               IF NOT #statIsArrayFieldClosed THEN
                 //field wasn't close as no deeper hierarchy exist, therfore the normal close opeartion is invalid
                 //close now here
                 #statInfoToWrite := CONCAT(IN1 := CHAR_TO_STRING(#BRACES_CLOSE), IN2 := CHAR_TO_STRING(#COMMA));
                 #statStackIndex -= #DECREMENT_BY_ONE;
               ELSE //reset flag
                 #statIsArrayFieldClosed := FALSE;
               END_IF;
               //open object
               #statInfoToWrite := CONCAT(IN1 := #statInfoToWrite, IN2 := CHAR_TO_STRING(#BRACES_OPEN), IN3 := CHAR_TO_STRING(#WHITE_SPACE));
               //increase stack index and push closing elements on to it
               #statStackIndex += #INCREMENT_BY_ONE;
               #statStackIndexOpenElement[#statStackIndex] := #BRACES_CLOSE;
             END_IF;

             IF NOT (#statIsArrayOpen AND #statArrayName = #tree[#statIndexTreeArray].key)  THEN
               //write key not in case array is open and key is the same array name
               //this indicates simple array structure e.g "ArrayName":["ArrayValue1","ArrayValue2"]
               //write key -> "key":
               #statInfoToWrite := CONCAT(IN1 := #statInfoToWrite, IN2 := CHAR_TO_STRING(#QUTATIONMARK),
                                          IN3 := #tree[#statIndexTreeArray].key, IN4 := CHAR_TO_STRING(#QUTATIONMARK),
                                          IN5 := CHAR_TO_STRING(#COLON), IN6 := CHAR_TO_STRING(#WHITE_SPACE));

             END_IF;

             //Move to state Write
             #statFbState := #FB_STATE_WRITE_TO_JSON;
             //Set state, that should be executed after writing
             //move on to next state
             #statFbNextState := #FB_STATE_VALUE_TYPE;

           END_REGION NEXT_ELEMENT 

         #FB_STATE_VALUE_TYPE: // Depending on value type, write value
           REGION VALUE DEPENDECY OF TYPE
             CASE #tree[#statIndexTreeArray].type OF

               #OBJECT:
                 REGION OBJECT
                   //nothing to do when type is object just add line feed, { openning will occur with next depth
                   #statInfoToWrite := CONCAT(IN1 := #statInfoToWrite, IN2 := CHAR_TO_STRING(#BRACES_OPEN));
                   //increase stack index and push closing elements on to it
                   #statStackIndex += #INCREMENT_BY_ONE;
                   #statStackIndexOpenElement[#statStackIndex] := #BRACES_CLOSE;
                 END_REGION OBJECT

               #ARRAY:
                 REGION ARRAY

                   IF (NOT #statIsArrayOpen) THEN
                     #statIsFirstElement := TRUE;
                     #statIsArrayOpen := TRUE;
                     //set Name of Array
                     #statArrayName := #tree[#statIndexTreeArray].key;

                     #statInfoToWrite := CONCAT(IN1 := CHAR_TO_STRING(#BRACKETS_OPEN), IN2 := CHAR_TO_STRING(#WHITE_SPACE));
                     //increase stack index and push closing elements on to it
                     #statStackIndex += #INCREMENT_BY_ONE;
                     #statStackIndexOpenElement[#statStackIndex] := #BRACKETS_CLOSE;

                     //case for underlaying object structure in array, prevent depth of simple array to have leading {
                     //simple array always has arrayname as key
                     IF #tree[#statIndexTreeArray].depth < #tree[#statIndexTreeArray + #NEXT_INDEX].depth
                       AND #tree[#statIndexTreeArray+ #NEXT_INDEX].key <> #statArrayName THEN
                       //open object
                       #statInfoToWrite := CONCAT(IN1 := #statInfoToWrite, IN2 := CHAR_TO_STRING(#BRACES_OPEN));
                       //increase stack index and push closing elements on to it
                       #statStackIndex += #INCREMENT_BY_ONE;
                       #statStackIndexOpenElement[#statStackIndex] := #BRACES_CLOSE;
                     END_IF;

                   END_IF;

                   // //null indicating that it is array definition, array information is written sepe
                   // //otherwise write value as string - value enclosed with quotation mark 
                   // IF(#tree[#statIndexTreeArray].value <> #NULL) THEN
                   //   #statInfoToWrite := CONCAT(IN1 := #statInfoToWrite, IN2 := CHAR_TO_STRING(#QUTATIONMARK),
                   //                              IN3 := #tree[#statIndexTreeArray].value, IN4 := CHAR_TO_STRING(#QUTATIONMARK));
                   // END_IF;
                 END_REGION ARRAY 

               #STRING:
                 REGION STRING

                   //wirte value as string - value enclosed with quotation mark 
                   IF (#tree[#statIndexTreeArray].value <> #NULL) THEN
                     #statInfoToWrite := CONCAT(IN1 := #statInfoToWrite, IN2 := CHAR_TO_STRING(#QUTATIONMARK),
                                                IN3 := #tree[#statIndexTreeArray].value, IN4 := CHAR_TO_STRING(#QUTATIONMARK));

                   ELSE // empty value still needs "" otherwise syntax error
                     #statInfoToWrite := CONCAT(IN1 := #statInfoToWrite, IN2 := CHAR_TO_STRING(#QUTATIONMARK),
                                                IN3 := CHAR_TO_STRING(#QUTATIONMARK));
                   END_IF;
                 END_REGION STRING

               #NUMBER, #BOOLEAN:
                 REGION NUMBER_BOOLEAN
                   //wirte value as number or boolean - value enclosed without quotation mark 
                   IF (#tree[#statIndexTreeArray].value <> #NULL) THEN
                     #statInfoToWrite := CONCAT(IN1 := #statInfoToWrite,
                                                IN2 := #tree[#statIndexTreeArray].value);
                   END_IF;
                 END_REGION NUMBER_BOOLEAN

               ELSE // Undefined state in state machine reached
                 REGION UNDEFINED STATE
                   #statStatus := #ERR_UNDEFINED_STATE;
                 END_REGION UNDEFINED STATE          

             END_CASE;

             //Move to state Write
             #statFbState := #FB_STATE_WRITE_TO_JSON;

             //Set state, that should be executed after writing
             //move on to next state
             #statFbNextState := #FB_STATE_NEXT_ELEMENT;

             IF #statIsLastElement OR #tree[#statIndexTreeArray].depth > #tree[#statIndexTreeArray + #NEXT_INDEX].depth THEN
               //Next Element has lower depth, therefore Elements have to be closed
               #statFbNextState := #FB_STATE_CLOSE_STACK_ELEMENT;
             ELSIF #statIsLastElement OR #tree[#statIndexTreeArray].depth = #tree[#statIndexTreeArray + #NEXT_INDEX].depth AND  NOT #statIsFirstElement THEN
                #statInfoToWrite := CONCAT(IN1 := #statInfoToWrite,
                                           IN2 := CHAR_TO_STRING(#COMMA));
             END_IF;
             //#statInfoToWrite := CONCAT(IN1 := #statInfoToWrite, IN2 := CHAR_TO_STRING(#LINE_FEED));



             //increase tree index to access next element 
             #statIndexTreeArray += #INCREMENT_BY_ONE;

           END_REGION VALUE DEPENDECY OF TYPE

         #FB_STATE_WRITE_TO_JSON: // Write to Byte Array
           REGION WRITE TO JSON                
             //add information to json byte array
             IF ((INT_TO_UINT(LEN(#statInfoToWrite)) + #statIndexJsonByteArray) < #statJsonByteLen) THEN
               Strg_TO_Chars(Strg := #statInfoToWrite,
                             pChars := #statIndexJsonByteArray,
                             Cnt => #tempCntCharsAdded,
                             Chars := #jsonByteArray);


               #statInfoToWrite := #EMPTY;
               //move index of byte array 
               #statIndexJsonByteArray += #tempCntCharsAdded;
               //move to next state previously allocated
               #statFbState := #statFbNextState;
             ELSE // Error: Index out of bounds
               #statStatus := #ERR_JSON_OUT_OF_BOUNDS;
             END_IF;

             IF #statLastElementIsClosed THEN
               //writer has written last information and execution is done
               #statStatus := #STATUS_EXECUTION_FINISHED;
               //current index equals count/size of json byte array
               #statCount := #statIndexJsonByteArray;
             END_IF;
           END_REGION WRITE TO JSON

         #FB_STATE_CLOSE_STACK_ELEMENT: //Close Open Stack Elements
           REGION CLOSE ELEMENT FROM STACK
             //close element with syntax </key>

             IF #statStackIndex >= 0 THEN //more open elements available, not all elements are closed

               //statInfoToWrite --> } or ]
               #statInfoToWrite := CHAR_TO_STRING(#statStackIndexOpenElement[#statStackIndex]);

               IF #statInfoToWrite = #BRACKETS_CLOSE THEN
                 //reset flag
                 #statIsArrayOpen := FALSE;

                 //first array key is used to recognize,
                 //beginning of new array field reset here, so it can be check for emptiness
                 #statFirstArrayKey := '';
               END_IF;

               //pop element from stack 
               #statStackIndex -= SINT_TO_INT(#DECREMENT_BY_ONE);

               IF #statStackIndex >= 0 THEN //more open elements available, not all elements are closed
                 //look at current stack item depth, if next tree element has 
                 IF NOT #statIsLastElement AND #statStackIndex = #tree[#statIndexTreeArray].depth THEN
                   //move to next element
                   //write comma as JSON dictates same depth a divided by comma,
                   //here we move on to the next elment with the same depth
                   #statInfoToWrite := CONCAT(IN1:=  #statInfoToWrite, IN2:= CHAR_TO_STRING(#COMMA));

                   // //if Array is still open and the same lenght is reached,
                   // //new element in array, distinguish new entry with BRACES
                   IF #statIsArrayOpen THEN
                     #statInfoToWrite := CONCAT(IN1 := #statInfoToWrite, IN2 := CHAR_TO_STRING(#BRACES_CLOSE), IN3 := CHAR_TO_STRING(#COMMA));
                     //pop element from stack 
                     #statStackIndex -= SINT_TO_INT(#DECREMENT_BY_ONE);
                     #statIsArrayFieldClosed := TRUE;
                   //   #statInfoToWrite := CONCAT(IN1 := #statInfoToWrite, IN2 := CHAR_TO_STRING(#BRACES_OPEN));
                   //   //increase stack index and push closing elements on to it
                   //   #statStackIndex += #INCREMENT_BY_ONE;
                   //   #statStackIndexOpenElement[#statStackIndex] := #BRACES_CLOSE;
                   END_IF;
                   #statFbNextState := #FB_STATE_NEXT_ELEMENT;

                 ELSE
                   //do nothing and return to fb state close element 
                   #statFbNextState := #FB_STATE_CLOSE_STACK_ELEMENT;
                 END_IF;

               ELSE
                 //no more open Elements, last Element was closed
                 #statIsLastElement := TRUE;

                 //only if this flag is set, can writer be finished
                 #statLastElementIsClosed := TRUE;

               END_IF;

             ELSE
               //no more open Elements, last Element was closed
               #statIsLastElement := TRUE;

               //only if this flag is set, can writer be finished
               #statLastElementIsClosed := TRUE;

             END_IF;
             //Move to state Write
             #statFbState := #FB_STATE_WRITE_TO_JSON;

           END_REGION CLOSE ELEMENT FROM STACK

         ELSE // Undefined state in state machine reached
           REGION UNDEFINED STATE
             #statStatus := #ERR_UNDEFINED_STATE;
           END_REGION UNDEFINED STATE     

       END_CASE;
       //Leave state machine if one of the following condition is true
       //1. state has not changed
       //2. error has occured
       //3. watchdog timer expired 
       //4. execution has finished
       // otherwise stay in state machine
     UNTIL (#statFbPreviousState = #statFbState OR #statStatus.%X15
       OR #instWatchdog.Q OR #statStatus = #STATUS_EXECUTION_FINISHED)
     END_REPEAT;
   END_REGION STATE_MACHINE

   REGION OUTPUTS
     // Write outputs
     IF (#statStatus = #STATUS_EXECUTION_FINISHED) AND (#statDone = FALSE) THEN // Execution finished without errors
       REGION EXECUTION FINSIHED
         #statDone := TRUE;
         #statBusy := FALSE;
         #statError := FALSE;
         // execution aborted --> set state no processing
         #statFbState := #FB_STATE_NO_PROCESSING;
       END_REGION EXECUTION FINSIHED

     ELSIF (#statStatus.%X15 = TRUE) AND (#statError = FALSE) THEN // Error occurred (#statStatus is 16#8000 to 16#FFFF)
       REGION ERROR OCCURED
         #statDone := FALSE;
         #statBusy := FALSE;
         #statError := TRUE;
         // execution aborted --> set state no processing
         #statFbState := #FB_STATE_NO_PROCESSING;
       END_REGION ERROR OCCURED

     ELSIF (#tempExecute = FALSE) AND ((#statDone = TRUE) OR (#statError = TRUE)) THEN // Reset outputs
       REGION EXECUTE RESETTED
         #statDone := FALSE;
         #statBusy := FALSE;
         #statError := FALSE;
         #statStatus := #STATUS_NO_CALL;
         // Reset application specific outputs
         #statCount := 0;
       END_REGION EXECUTE RESETTED
     END_IF;

     REGION WRITE STATIC VALUES TO OUTPUTS
       #done := #statDone;
       #busy := #statBusy;
       #error := #statError;
       #status := #statStatus;
       //  ENO mechanism is not used 
       ENO := TRUE;
       // Write application specific static values to outputs
       #count := #statCount;
     END_REGION WRITE STATIC VALUES TO OUTPUTS
   END_REGION OUTPUTS
END_FUNCTION_BLOCK

// folder: LStream/Utilities

FUNCTION "LStream_FindStringInByteCharArrayAdv" : DInt   // FC2, SCL
TITLE = LStream_FindStringInCharArrayAdv
{ S7_Optimized_Access := 'TRUE' }
AUTHOR : DI_FA_S_SUP_EuC
FAMILY : LStream
VERSION : 1.0
// Finds string in char array
   VAR_INPUT
      searchFor : String;   // Text that is searched for
      startPosition : DInt;   // Start position in array
   END_VAR
   VAR_IN_OUT
      searchIn : Array[*] of Byte;   // Array of Char to search in
   END_VAR
   VAR_TEMP
      tempLowerBound : DInt;   // Lower bound of given array
      tempNumElements : UDInt;   // Number of elements in given array
      tempLenSearchFor : Int;   // Length of text that is seached for
      tempPosInArray : DInt;   // Position in array during search (0-based)
      tempPosInString : Int;   // Position in working string during search
      tempString : String;   // Temporary string to work with
   END_VAR
   // Ret_Val : Returns the index of found string
   VAR CONSTANT
      FIRST_DIM : USInt := 1;   // Constant for first array dimenson
      MAX_LEN_STRING : UInt := 254;   // Max. length of String
   END_VAR
BEGIN
   REGION BLOCK INFO HEADER
     //===============================================================================
     // SIEMENS AG / (c)Copyright 2021
     //-------------------------------------------------------------------------------
     // Title:            LStream_FindStringInByteCharArrayAdv
     // Comment/Function: Searches for a specified string within an array of char
     // Library/Family:   LStream
     // Author:           DI FA S SUP E&C
     // Tested with:      S7-1500 V2.8
     // Engineering:      TIA Portal V16
     // Restrictions:     --
     // Requirements:     --
     //-------------------------------------------------------------------------------
     // Change log table:
     // Version  | Date       | Expert in charge | Changes applied
     //----------|------------|------------------|------------------------------------
     // 01.00.00 | 2021-03-10 |DI FA S SUP E&C   | First released version
     //===============================================================================
   END_REGION

   // Initialization
   #tempPosInString := 0;
   #tempPosInArray := #startPosition;
   #tempLenSearchFor := LEN(#searchFor);
   #LStream_FindStringInByteCharArrayAdv := -1;

   // Get number of elements
   #tempLowerBound := LOWER_BOUND(ARR := #searchIn, DIM := #FIRST_DIM);
   #tempNumElements := DINT_TO_UDINT(UPPER_BOUND(ARR := #searchIn, DIM := #FIRST_DIM) - #tempLowerBound + 1);

   IF (#tempPosInArray > #tempNumElements) THEN
       RETURN;
   END_IF;

   // Search for beginning of text until something was found and
   // as long as the index is less than the array size / number of elements in array
   WHILE ((#tempPosInString <= 0) AND (#tempPosInArray < #tempNumElements)) DO
       // Convert Chars to String
       Chars_TO_Strg(Chars := #searchIn,
                     pChars := #tempPosInArray,
                     Cnt := UDINT_TO_UINT(MIN(IN1 := #MAX_LEN_STRING, IN2 := #tempNumElements)),
                     Strg => #tempString);

       // Search for text at beginning
       #tempPosInString := FIND(IN1 := #tempString, IN2 := #searchFor);

       // Keyword was found
       IF #tempPosInString > 0 THEN
           // Output position of string
           #LStream_FindStringInByteCharArrayAdv := #tempLowerBound + #tempPosInArray + #tempPosInString - 1;
           EXIT;
       ELSE
           // Otherwise continue search in next string minus length of text at beginning to ensure
           // keywords are not broken up at the end of a string and thus missed
           #tempPosInArray += UINT_TO_INT(#MAX_LEN_STRING) - #tempLenSearchFor;
       END_IF;
   END_WHILE;
END_FUNCTION

// ===== library types =====

// folder: LMQTT

TYPE "LMQTT_typeConnParam"
TITLE = LMQTT_typeConnParams
// Specifies connection parameters for the mqtt connection
   STRUCT
      hwId : Hw_Any;   // Hardware identifier of the interface. 0: interface is selected automatically
      connId : Conn_Ouc;   // Unique connection identifier
      brokerAddress : Struct   // Information on the MQTT broker
         qdnAddress : String;   // Fully qualified domain name of the broker. must end with a dot "."
         ipAddress : IP_V4;   // If no FQDN is used, enter ip-address of the broker instead
         port : UInt;   // Enter the port of the mqtt broker
      END_STRUCT;
      tls : Struct   // Parameters for TLS encryption
         enableTls : Bool;   // TRUE: Enables TLS, FALSE: disable TLS
         validateServerIdentity : Bool;   // TRUE: Validate server certificate, FALSE: No validation of server certificate
         brokerCert : UDInt;   // ID of the broker's certificate in TIA Portal
         clientCert : UDInt;   // ID of the client's certificate in TIA Portal
      END_STRUCT;
      keepAlive : UInt;   // Keepalive mechanism for MQTT in seconds. 0: disabled.
   END_STRUCT;
END_TYPE

(* ===== HMI "HMI_RT_1" =====
system functions are stored by id; their names below are inferred from use
connection "HMI_Conexión_1": ETHERNET, SMART_S7_1500_OMS

HMI tags "VariablesHMI"
   "MqttSubscribe" : Bool = PLC MqttDB.control.subscribe, 1 s
   "JsonDeserialize" : Bool = PLC JSON_DeserializParamDB.execute, 1 s
   "JsonSerialize" : Bool = PLC JSON_SerializParamDB.execute AT %M1.2, 1 s
   "MqttConnect" : Bool = PLC MqttDB.control.connect AT %DB1.DBX0.0, 1 s
   "MqttConnected" : Bool = PLC MqttConnected AT %M1.0, 1 s
   "MqttDataReceived" : Bool = PLC MqttDataReceived AT %M1.1, 1 s
   "MqttPublish" : Bool = PLC MqttDB.control.publish AT %M1.2, 1 s
   "MqttSubscribed" : Bool = PLC MqttSubscribed AT %M1.3, 1 s
   "MqttUnsubscribed" : Bool = PLC MqttUnsuscribed AT %M1.4, 1 s
   "No_of_Items" : USInt = PLC AASassetDB.Agent2PLC.Operation.No_of_Items, 1 s
   "Service_Type" : UDInt = PLC AASassetDB.Agent2PLC.Operation.Ref_Service_Type AT %DB1.DBD0, 1 s
   "Item_Number" : USInt = PLC AASassetDB.PLC2Agent.Id.Item_Number AT %DB1.DBB0, 1 s
   "Item_Completed" : Bool = PLC AASassetDB.Control.Flag_Item_Completed AT %DB1.DBX0.0, 1 s
   "Service_Completed" : Bool = PLC AASassetDB.Control.Flag_Service_Completed AT %DB1.DBX0.0, 1 s
   "MqttUnsuscribe" : Bool = PLC MqttDB.control.unsubscribe AT %DB1.DBX0.0, 1 s
   "New_Service" : Bool = PLC AASassetDB.Control.Flag_New_Service AT %DB1.DBX0.0, 1 s
   "Initial_Time" : LDT = PLC AASassetDB.PLC2Agent.Data.Initial_Time_Stamp AT %DB1.DBX0.0, 1 s
   "Final_Time" : LDT = PLC AASassetDB.PLC2Agent.Data.Final_Time_Stamp AT %DB1.DBX0.0, 1 s
   "Service_Time" : LDT = PLC AASassetDB.PLC2Agent.Data.Service_Time_Stamp AT %DB1.DBX0.0, 1 s

Template "Plantilla_1" 1280x800
   Button "Salir" at 1182,752 size 67x47; TextOff 'Salir'; PictureOff "ExitRuntime_KTP1200_Basic_PN_TR"; PictureOn "ExitRuntime_KTP1200_Basic_PN_TR"
      on Release: StopRuntime(0)
   Button "Template_Button" at 1054,752 size 67x47; TextOff 'Text'
   Button "Template_Button_1" at 926,752 size 67x47; TextOff 'Text'
   Button "Template_Button_2" at 798,752 size 67x47; TextOff 'Text'
   Button "Template_Button_3" at 670,752 size 67x47; TextOff 'Text'
   Button "Template_Button_4" at 542,752 size 67x47; TextOff 'Text'
   Button "Template_Button_5" at 414,752 size 67x47; TextOff 'Text'
   Button "Template_Button_6" at 286,752 size 67x47; TextOff 'Text'
   Button "Template_Button_7" at 158,752 size 67x47; TextOff 'Text'
   Button "Imagen inicial" at 30,752 size 67x47; TextOff 'Imagen inicial'; PictureOff "NavigateHome_KTP1200_Basic_PN_TR"; PictureOn "NavigateHome_KTP1200_Basic_PN_TR"
      on Release: ActivateScreen("Imagen raíz", 0)

screen "Imagen raíz" 1280x800, template "Plantilla_1"
   Switch "Interruptor_1" at 305,215 size 66x26; TextOn 'OFF'; CaptionText 'Switch'; TextOff 'ON'
      on SwitchOff: ResetBit("MqttConnect")
      on SwitchOn: SetBit("MqttConnect")
   TextField "Campo de texto_1" at 43,213 size 244x29; Text 'Conexión con el bróker'
   TextField "Campo de texto_5" at 43,253 size 224x29; Text 'Suscripción al bróker'
   TextField "Campo de texto_6" at 45,523 size 163x29; Text 'Dato publicado'
   Circle "Círculo_3" at 387,213 size 29x29
      Appearance <- "MqttConnected"
   TextField "Campo de texto_16" at 43,297 size 273x29; Text 'Datos recibidos de broker'
   Circle "Círculo_8" at 387,297 size 29x29
      Appearance <- "MqttDataReceived"
   TextField "Campo de texto_17" at 43,326 size 194x29; Text 'Deserializar datos'
   Button "Botón_2" at 297,332 size 82x32; TextOff 'deserial'
      on Release: ResetBit("JsonDeserialize")
      on Press: SetBit("JsonDeserialize")
   Switch "Interruptor_2" at 305,255 size 66x26; TextOn 'OFF'; CaptionText 'Switch'; TextOff 'ON'
      on SwitchOn: SetBit("MqttSubscribe"); ResetBit("MqttUnsuscribe")
      on SwitchOff: ResetBit("MqttSubscribe"); SetBit("MqttUnsuscribe")
   Circle "Círculo_2" at 387,253 size 29x29
      Appearance <- "MqttSubscribed"
   TextField "Campo de texto_2" at 45,486 size 175x29; Text 'Dato serializado'
   IOField "Campo ES_1" at 816,228 size 68x32; FormatPattern 99
      ProcessValue <- "Service_Type"
   IOField "Campo ES_2" at 955,228 size 68x32; FormatPattern 99
      ProcessValue <- "No_of_Items"
   TextField "Campo de texto_7" at 944,193 size 89x29; Text 'Nº Item'
   TextField "Campo de texto_3" at 806,193 size 87x29; Text 'Servicio'
   IOField "Campo ES_3" at 726,427 size 68x32; FormatPattern 99
      ProcessValue <- "Item_Number"
   TextField "Campo de texto_8" at 673,398 size 174x29; Text 'Item Completed'
   Circle "Círculo_1" at 887,398 size 29x29
      Appearance <- "Item_Completed"
   TextField "Campo de texto_9" at 673,472 size 198x29; Text 'Service Completed'
   Circle "Círculo_4" at 887,472 size 29x29
      Appearance <- "Service_Completed"
   TextField "Campo de texto_10" at 673,360 size 133x29; Text 'New Service'
   Circle "Círculo_5" at 887,360 size 29x29
      Appearance <- "New_Service"
   Circle "Círculo_6" at 389,489 size 29x29
      Appearance <- "JsonSerialize"
   Circle "Círculo_7" at 389,529 size 29x29
      Appearance <- "MqttPublish"
   TextField "Campo de texto_4" at 667,544 size 199x29; Text 'Initial Time Stamp'
   TextField "Campo de texto_11" at 670,598 size 186x29; Text 'Final Time Stamp'
   TextField "Campo de texto_12" at 670,652 size 211x29; Text 'Service Time Stamp'
   TextField "Campo de texto_13" at 831,301 size 207x47; Text 'Producción'
   TextField "Campo de texto_14" at 831,134 size 163x47; Text 'Solicitud'
   TextField "Campo de texto_15" at 128,143 size 214x47; Text 'Suscripción'
   TextField "Campo de texto_18" at 130,425 size 213x47; Text 'Publicación'
   TextField "Campo de texto_19" at 327,19 size 640x66; Text 'Célula robotizada - UR3e'
   IOField "Campo ES_4" at 968,539 size 209x39; FormatPattern 9999999999999999999999999999999999999999
      ProcessValue <- "Initial_Time"
   IOField "Campo ES_5" at 968,593 size 209x39; FormatPattern 9999999999999999999999999999999999999999
      ProcessValue <- "Final_Time"
   IOField "Campo ES_6" at 968,647 size 209x39; FormatPattern 9999999999999999999999999999999999999999
      ProcessValue <- "Service_Time"
*)